// TIA Portal project "THELMA3_200224" (V15.1) (continued)
               #SDataDummy := CONCAT(IN1 := #SDataDummy, IN2 := 'BBD');
               #SDataDummy := CONCAT(IN1 := #SDataDummy, IN2 := #ExtDate);
               Strg_TO_Chars(Strg := #SDataDummy,
                             pChars := 1,
                             Cnt => #Dummy2,
                             Chars := #SData);
               #SData[15 + #LenDummy] := #End;
               #SLen := 15 + #LenDummy + 1;
               #RLen := 3;
               #Step := 0;
               #STrig := TRUE;
               #RdataTime := FALSE;
               #RdataAlarm := FALSE;
               #RdataBatch := FALSE;
               #RdataBBD := TRUE;
               #RdataLabel := FALSE;
               #Selected := FALSE;
           ELSIF #MarketRegCode <> '' AND #ExtDate <> '' THEN // print all on the second row
               #CommandHead := 'U'; //head for update user field
               #LenDummy := LEN(#MarketRegCode);
               #SDataDummy := CONCAT(IN1 := #CommandHead, IN2 := #SecondField);
               #SDataDummy := CONCAT(IN1 := #SDataDummy, IN2 := #NewLine);
               #SDataDummy := CONCAT(IN1 := #SDataDummy, IN2 := #MarketRegCode);
               #SDataDummy := CONCAT(IN1 := #SDataDummy, IN2 := 'BBD');
               #SDataDummy := CONCAT(IN1 := #SDataDummy, IN2 := #ExtDate);
               Strg_TO_Chars(Strg := #SDataDummy,
                             pChars := 1,
                             Cnt => #Dummy2,
                             Chars := #SData);
               #SData[21 + #LenDummy] := #End;
               #SLen := 21 + #LenDummy + 1;
               #RLen := 3;
               #Step := 0;
               #STrig := TRUE;
               #RdataTime := FALSE;
               #RdataAlarm := FALSE;
               #RdataBatch := FALSE;
               #RdataBBD := TRUE;
               #RdataLabel := FALSE;
               #Selected := FALSE;
           END_IF;
       ELSIF #Step =5 THEN
           //command for selecting the label
           #CommandHead := 'M'; //head for current status of the printer
           #SData[0] := #Start;
           IF #MDR_Flag = TRUE THEN //select the MDR layout 
               #SDataDummy := CONCAT(IN1 := #CommandHead, IN2 := #MDR_LabelName);
               Strg_TO_Chars(Strg := #SDataDummy,
                             pChars := 1,
                             Cnt => #Dummy2,
                             Chars := #SData);
               #SData[5] := #End;
               #RLen := 3;
               #SLen := 6;
           ELSE
               #LenLabel := LEN(#NMDR_LabelName);
               #SDataDummy := CONCAT(IN1 := #CommandHead, IN2 := #NMDR_LabelName);
               Strg_TO_Chars(Strg := #SDataDummy,
                             pChars := 1,
                             Cnt => #Dummy2,
                             Chars := #SData);
               #SData[2+#LenLabel] := #End;
               #RLen := 3;
               #SLen := 3+#LenLabel;
           END_IF;
           #STrig := TRUE;
           #Step := 0;
           #RdataAlarm := FALSE;
           #RdataTime := FALSE;
           #RdataBatch := FALSE;
           #RdataBBD := FALSE;
           #RdataLabel := TRUE;
       ELSE
           #STrig := FALSE;
       END_IF;
   END_REGION

   REGION Feedback
       // Statement section REGION
       //Expect to receive "ACT"
       IF #DataReceived = TRUE THEN
           #StartTNR := FALSE;
           IF #RdataTime = TRUE THEN //check for the feedback for the time command
               FOR #i := 0 TO 56 DO
                   #TimeReceivedData[#i] := #RData[#i];
               END_FOR;
               IF #TimeReceivedData[0] = 16#24 THEN
                   #TimeOK := TRUE;
                   #TimeReceivedData[0] := 16#30;//clear the buffer
               ELSE
                   #TimeOK := FALSE;
               END_IF;
               #RdataTime := FALSE;
           ELSIF #RdataAlarm = TRUE THEN//check for the feedback for the alarm command
               FOR #i := 0 TO 56 DO
                   #AlarmReceivedData[#i] := #RData[#i];
               END_FOR;
               IF #AlarmReceivedData[7] = 16#30  THEN
                   #AlarmCheck := TRUE;

                   FOR #i := 0 TO 8 DO
                       #PrinterAlarmStatus[#i] := #AlarmReceivedData[#i];//save the status data for processing
                   END_FOR;
                   #AlarmReceivedData[7] := 16#31;//clear the buffer
               ELSE
                   #AlarmCheck := FALSE;
               END_IF;
               #RdataAlarm := FALSE;
           ELSIF #RdataBatch = TRUE THEN//check for the feedback for the buffer command
               FOR #i := 0 TO 56 DO
                   #BatchReceivedData[#i] := #RData[#i];
               END_FOR;
               IF #BatchReceivedData[0] = 16#24 THEN
                   #BatchOK := TRUE;
                   #BatchReceivedData[0] := 16#30;//clear the buffer
               ELSE
                   #BatchOK := FALSE;
               END_IF;
               #RdataBatch := FALSE;
           ELSIF #RdataBBD = TRUE THEN//check for the feedback for the buffer command
               FOR #i := 0 TO 56 DO
                   #BBD_ReceivedData[#i] := #RData[#i];
               END_FOR;
               IF #BBD_ReceivedData[0] = 16#24 THEN
                   #BBD_OK := TRUE;
                   #BBD_ReceivedData[0] := 16#30;//clear the buffer
               ELSE
                   #BBD_OK := FALSE;
               END_IF;
               #RdataBBD := FALSE;
           ELSIF #RdataLabel = TRUE THEN//check for the feedback for the buffer command
               FOR #i := 0 TO 56 DO
                   #LabelReceivedData[#i] := #RData[#i];
               END_FOR;
               IF #LabelReceivedData[0] = 16#24 THEN
                   #LabelOK := TRUE;
                   #LabelReceivedData[0] := 16#30;//clear the buffer
               ELSE
                   #LabelOK := FALSE;
               END_IF;
               #RdataLabel := FALSE;
           END_IF;
       ELSIF #DataSent = TRUE THEN // command send noting received
           #StartTNR := TRUE;
           IF #RdataTime = TRUE THEN
               #TimeOK := FALSE;
           END_IF;
           IF #RdataAlarm = TRUE THEN
               #AlarmCheck := FALSE;
           END_IF;
           IF #RdataBatch = TRUE THEN
               #BatchOK := FALSE;
           END_IF;
           IF #RdataBBD = TRUE THEN
               #BBD_OK := FALSE;
           END_IF;
           IF #RdataLabel = TRUE THEN
               #LabelOK := FALSE;
           END_IF;
       END_IF;
   END_REGION

   REGION Sending
       // Send the batch number when it is changed or for reconnection
       #SelectingR(CLK:=#LabelSelecting);
       #ReconnectR(CLK := #ConnectionStatus);
       #MDR_R(CLK := #MDR_Flag);
       #MDR_F(CLK := #MDR_Flag);
       #BlockedR(CLK := #BlockedProduct);
       #BlockedF(CLK := #BlockedProduct);
       //select the label
       IF #MDR_F.Q = TRUE OR #MDR_R.Q = TRUE OR #SelectingR.Q = TRUE OR #ReconnectR.Q = TRUE OR #NLabelChanged = TRUE THEN
           #Step := 5; //selecting the label
           IF #MDR_Flag = TRUE THEN
               #Selected := TRUE; //send the first row
               #First := TRUE;////send the second row
           END_IF;
       END_IF;
       // set the step to 3 after label is selected (small delay to make sure that the label is loaded)
       #BatchAfterLabelT(IN := #Selected,
                         PT := T#2S);
       IF #BatchAfterLabelT.Q = TRUE THEN
           #Step := 3;
       END_IF;
       //send the update information
       // Send the updateble data when it is changed and step 4 is done
       IF (#PlainDataChanged = TRUE OR #BlockedR.Q = TRUE OR #BlockedF.Q = TRUE) AND #SelectingR.Q = FALSE THEN
           #Step := 3; //send plain data
           #Selected := FALSE;
           #First := TRUE;
       END_IF;
       //set the step to 4 after the first row is send
       #SecondAfterFirstT(IN:=#First,
                          PT:=T#4S);
       IF #SecondAfterFirstT.Q = TRUE THEN
           #Step := 4;
       END_IF;
       // Send time and alarm commands
       //every 10 minute synchronise time
       #TimeSynchT(IN := #TimeSynchEnable,
                  PT := #TimeSynchPeriod);
       IF #TimeSynchT.Q = TRUE THEN
           #Step := 1;
           #TimeSynchEnable := FALSE;
       ELSIF #ConnectionStatus = TRUE AND NOT (#MDR_F.Q= TRUE OR #MDR_R.Q =TRUE OR #SelectingR.Q = TRUE OR #ReconnectR.Q = TRUE OR #NLabelChanged = TRUE) AND NOT (#PlainDataChanged = TRUE OR #BlockedR.Q = TRUE OR #BlockedF.Q = TRUE) THEN
           #TimeSynchEnable := TRUE;
       ELSE
           #TimeSynchEnable := FALSE;
       END_IF;
       //every 5 minute check for alarm
       #AlarmCheckT(IN := #AlarmCheckEnable,
                   PT := #AlarmCheckPeriod + T#20MS);//+20ms to avoid conflict
       IF #AlarmCheckT.Q = TRUE THEN
           #Step := 2;
           #AlarmCheckEnable := FALSE;
       ELSIF #ConnectionStatus = TRUE AND NOT (#MDR_F.Q = TRUE OR #MDR_R.Q = TRUE OR #SelectingR.Q = TRUE OR #ReconnectR.Q = TRUE OR #NLabelChanged = TRUE) AND NOT(#PlainDataChanged = TRUE OR #BlockedR.Q = TRUE OR #BlockedF.Q = TRUE) THEN
           #AlarmCheckEnable := TRUE;
       ELSE
           #AlarmCheckEnable := FALSE;
       END_IF;
   END_REGION

   REGION send try
       //if not receiving feedback after 10ms send a commad again
       #NotReceiveT(IN := #StartTNR,
                   PT := #TimeNR,
                   Q => #SendAgainTrigger);
       IF #SendAgainTrigger = TRUE THEN
           #StartTNR := FALSE;
       END_IF;
   END_REGION
   (*
   REGION ConnReestablised
       // connection Re-Established Rotinue. It try 5 times to connect to the printer, if not succsess enable time out error
       #ConnAgainT(IN := #ReTry,
                  PT := T#5S);// time out for reconnection
       //try five times to connect
       #ConnTryCountC(CU := #ReTry,
                     R := #ConnectionStatus,
                     PV := 5,
                     Q => #TimeOutError);
   END_REGION
   *)
END_REGION
END_FUNCTION_BLOCK

FUNCTION_BLOCK "CON_PlainHandle"   // FB2, FBD
{ S7_Optimized_Access := 'TRUE' }
VERSION : 0.1
   VAR_INPUT
      Heartbeat : Bool;
      NewArtBaseFlag : String;
      NewMDR_Flag : String;
      NewBatchNum : String;
      NewArtBaseNum : UDInt;
      NewMarketRegCode : String;
      NewBBD : String;
   END_VAR
   VAR_OUTPUT
      Error : Bool;
      ActualBatchNumSTR : String;
      ActualArtBaseNumSTR : String;
      ActualMarketRegCodeSTR : String;
      ActualBBD_STR : String;
      HeartbeatToPlain : Bool;
   END_VAR
   VAR
      NewDataPlain : Bool;
      ActualMDR_FlagSTR : String;
      ActualArtBaseFlagSTR : String;
      ActualBatchNum : String;
      ActualArtBaseNum : UDInt;
      ActualMDR_Flag : Bool;
      ActualArtFlag : Bool;
      HeartbeatT : TON_TIME;
      PrintSecondRow : Bool;
      HeartbeatT_2 : TON_TIME;
      CountC : CTU_INT;
   END_VAR
   VAR_TEMP
      i : Int;
      NewBatchLen : UInt;
      Correction : Array[0..13] of Char;
      CorrectionSTR : String;
      TmpB1 : Bool;
      TmpB2 : Bool;
   END_VAR
   VAR CONSTANT
      BatchSize : UInt := 10;
   END_VAR
BEGIN

REGION Network 1 (SCL)
   REGION connection
       // check the heartbeat from MES-OPC
     #HeartbeatT(IN:=NOT(#Heartbeat),
                 PT:=T#30S);
     IF #HeartbeatT.Q = TRUE THEN
         #TmpB1 := TRUE;
       ELSE
           #TmpB1 := FALSE;
       END_IF;
       #HeartbeatT_2(IN:=#Heartbeat,
                     PT:=T#30S);
       IF #HeartbeatT_2.Q = TRUE THEN
           #TmpB2 := TRUE;
       ELSE
           #TmpB2 := FALSE;
       END_IF;
       IF #TmpB1 OR #TmpB2 THEN
           #Error := 1;
       ELSE
           #Error := 0;
       END_IF;

       //Send the Heartbeat to MES-OPC
       #CountC(CU:="Clock_1Hz",
               PV:=15,
               Q=>#HeartbeatToPlain);
       IF #CountC.CV > 29 THEN
           #CountC.CV := 0;
       END_IF;
   END_REGION
   REGION Flags
       // check for flags 
       IF #NewArtBaseFlag = 'Y' THEN
           #ActualArtFlag := TRUE;
       ELSE
           #ActualArtFlag := FALSE;
       END_IF;
       IF #NewMDR_Flag = 'Y' THEN
           #ActualMDR_Flag := TRUE;
       ELSE
           #ActualMDR_Flag := FALSE;
       END_IF;
   END_REGION

   REGION input changing
       // check for input number changing

       IF  #NewBatchNum <> #ActualBatchNum  OR  #NewArtBaseNum <> #ActualArtBaseNum OR #NewMarketRegCode <>#ActualMarketRegCodeSTR OR #NewBBD <> #ActualBBD_STR OR #NewArtBaseFlag <> #ActualArtBaseFlagSTR THEN
           #NewDataPlain := TRUE;
       ELSE
           #NewDataPlain := FALSE;
       END_IF;
       IF #NewBBD <> #ActualBBD_STR OR #NewMarketRegCode <> #ActualMarketRegCodeSTR THEN
           #PrintSecondRow := TRUE;
       ELSE
           #PrintSecondRow := FALSE;
       END_IF;
    //   IF #NewMDR_Flag <> #ActualMDR_FlagSTR THEN
    //       #MDR_FlagChange := TRUE;
   //    ELSE
   //        #MDR_FlagChange := FALSE;
   //    END_IF;
     //  IF #NewArtBaseFlag <> #ActualArtBaseFlagSTR THEN
     //      #ArtBaseFlagChange := TRUE;
     //  ELSE
    //       #ArtBaseFlagChange := FALSE;
    //   END_IF;
   END_REGION
   REGION assign plain data
       FOR #i := 0 TO 13 DO
           #Correction[#i] := '0';
       END_FOR;
       // Statement section REGION
       #ActualArtBaseNum := #NewArtBaseNum;
       #ActualMarketRegCodeSTR := #NewMarketRegCode;
       #ActualBatchNum := #NewBatchNum;
       #ActualBBD_STR := #NewBBD;
       #ActualMDR_FlagSTR := #NewMDR_Flag;
       #ActualArtBaseFlagSTR := #NewArtBaseFlag;
       //Actual Batch in 10 digits (3 factoryID+7 batch ID)
       #NewBatchLen := INT_TO_UINT(LEN(#NewBatchNum));
       IF #NewBatchLen < #BatchSize THEN
           Chars_TO_Strg(Chars := #Correction,
                         pChars := 0,
                         Cnt := (#BatchSize - #NewBatchLen),
                         Strg => #CorrectionSTR);
           #ActualBatchNumSTR := CONCAT(IN1 := #CorrectionSTR, IN2 := #NewBatchNum);
       ELSE
           #ActualBatchNumSTR := #NewBatchNum;
       END_IF;
     //Art base number
       VAL_STRG(IN := #NewArtBaseNum,
                SIZE := 0,
                PREC := 0,
                FORMAT := 0,
                P := 1,
                OUT => #ActualArtBaseNumSTR);
   END_REGION
END_REGION
END_FUNCTION_BLOCK

FUNCTION_BLOCK "ProgramReader"   // FB3, FBD
{ S7_Optimized_Access := 'TRUE' }
VERSION : 0.1
   VAR_INPUT
      Value : Array[0..9] of Char;
      MaterialNumber : UDInt;
      ReaderRead : Bool;
      ReaderNoRead : Bool;
      ExtTrigger : Bool;
      ResetFaults : Bool;
      ResetCounters : Bool;
   END_VAR
   VAR_OUTPUT
      Reading : UDInt;
      Msg_NoRead : Bool;
      Fault_MisMatch : Bool;
      Fault_NoRead : Bool;
      Fault_Trigger : Bool;
   END_VAR
   VAR_IN_OUT
      NumGross : UDInt;
      NumRead : UDInt;
      NumNoRead : UDInt;
      NumMatch : UDInt;
      NumNoMatch : UDInt;
   END_VAR
   VAR
      ReadingDInt : UDInt;
      ReadingSTR : String;
      MaterialNumberSTR : String;
      CompDINOut1 : Bool;
      HF_PosEdge1 : Bool;
      HF_PosEdge2 : Bool;
      HF_PosEdge3 : Bool;
      HF_PosEdge4 : Bool;
      HF_PosEdge5 : Bool;
      HF_PosEdge6 : Bool;
      HF_PosEdge7 : Bool;
      HF_PosEdge8 : Bool;
      HF_PosEdge9 : Bool;
      HF_NegEdge1 : Bool;
      HF_NegEdge2 : Bool;
      HF_MisMatch : Bool;
      HF_NoRead : Bool;
      HF_FltTrigger : Bool;
      HF_MisTrigger : Bool;
      HF_FltNoRead : Bool;
      T_FltNoRead : IEC_TIMER;
      Time_FltNoRead : Time := T#500MS;
      T_FltTriggerWatchdog : IEC_TIMER;
      Time_FltTriggerWatchdog : Time := T#5s;
   END_VAR
   VAR RETAIN
      C_FltNoRead : IEC_COUNTER;
      C_FltNoRead100 : IEC_COUNTER;
   END_VAR
   VAR
      TriggerCTR : "Counter_32Bit";
      ReadCTR : "Counter_32Bit";
      NoReadCTR : "Counter_32Bit";
      MatchCTR : "Counter_32Bit";
      NoMatchCTR : "Counter_32Bit";
      IEC_Timer_0_Instance : TP_TIME;
      MisTriggerCTR : "Counter_32Bit";
      NumMisTrigger : UDInt;
      NumNoReadGross : UDInt;
      EmptyBuffer : Bool;
      ReadData : Bool;
      DataValid : Bool;
      IEC_Timer_0_Instance_1 : TON_TIME;
   END_VAR
   VAR RETAIN
      Mis_3_row : CTU_INT;
   END_VAR
   VAR_TEMP   // added for the SCL form of the ladder/FBD networks
      _w1 : Bool;
   END_VAR
BEGIN

REGION Network 1
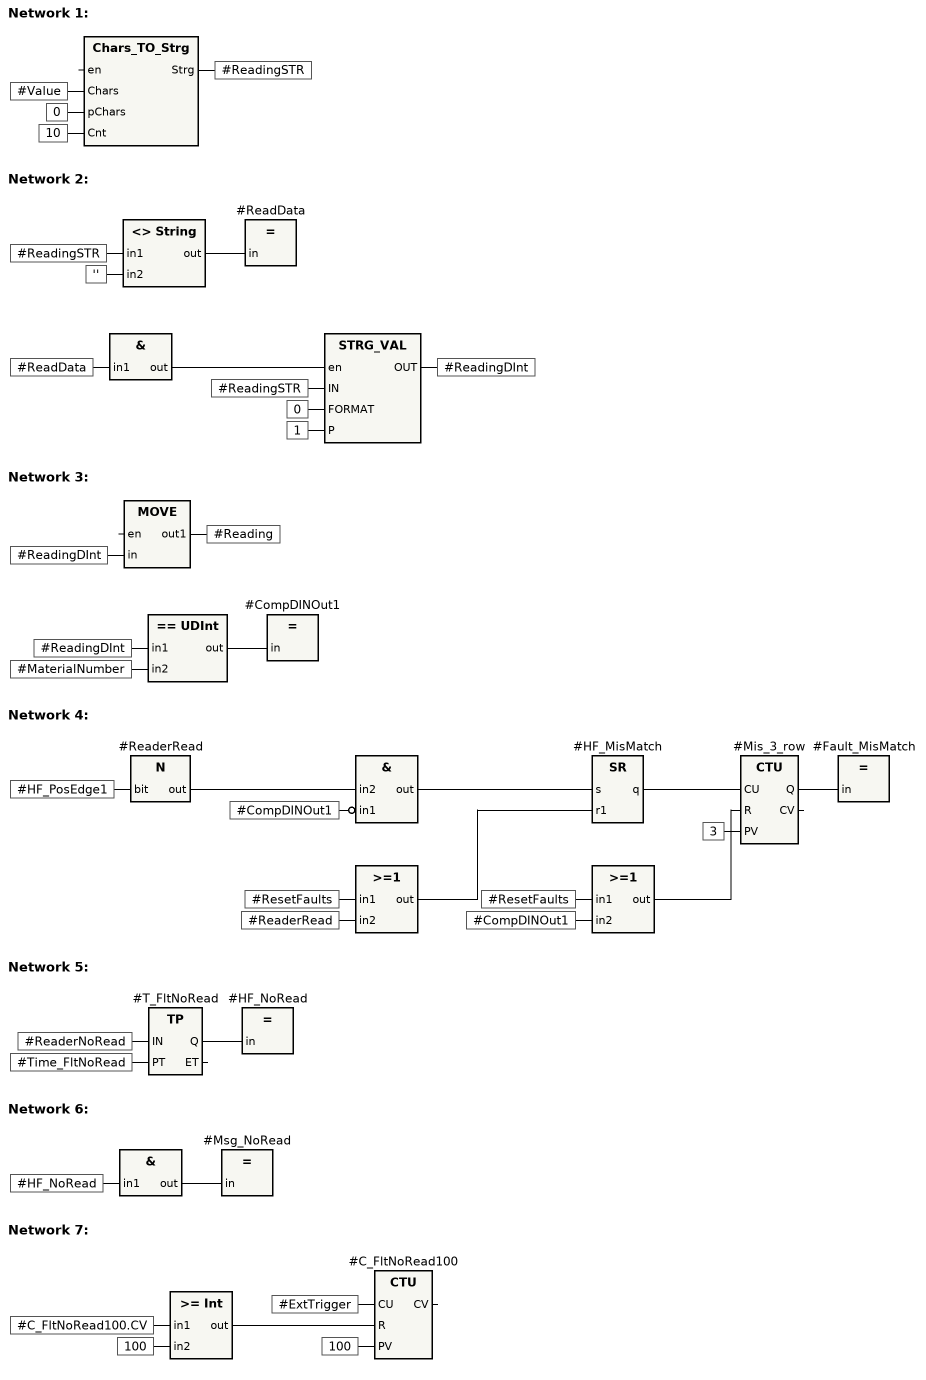
   // no SCL statement known for Chars_TO_Strg: written as a call
   Chars_TO_Strg(Chars := #Value, pChars := 0, Cnt := 10, Strg => #ReadingSTR);
END_REGION

REGION Network 2
   #ReadData := #ReadingSTR <> '';
   IF #ReadData THEN STRG_VAL(IN := #ReadingSTR, FORMAT := 0, P := 1, OUT => #ReadingDInt); END_IF;
END_REGION

REGION Network 3
   #Reading := #ReadingDInt;
   #CompDINOut1 := #ReadingDInt = #MaterialNumber;
END_REGION

REGION Network 4
   #_w1 := NOT #ReaderRead AND #HF_PosEdge1;   // falling edge of #ReaderRead
   #HF_PosEdge1 := #ReaderRead;
   IF #_w1 AND NOT #CompDINOut1 THEN
       #HF_MisMatch := TRUE;   // SR flip-flop
   END_IF;
   IF #ResetFaults OR #ReaderRead THEN #HF_MisMatch := FALSE; END_IF;
   #Mis_3_row(CU := #HF_MisMatch, R := #ResetFaults OR #CompDINOut1, PV := 3);   // CTU
   #Fault_MisMatch := #Mis_3_row.Q;
END_REGION

REGION Network 5
   #T_FltNoRead.TP(IN := #ReaderNoRead, PT := #Time_FltNoRead);
   #HF_NoRead := #T_FltNoRead.Q;
END_REGION

REGION Network 6
   #Msg_NoRead := #HF_NoRead;
END_REGION

REGION Network 7
   #C_FltNoRead100.CTU(CU := #ExtTrigger, R := #C_FltNoRead100.CV >= 100, PV := 100);
END_REGION

REGION Network 8
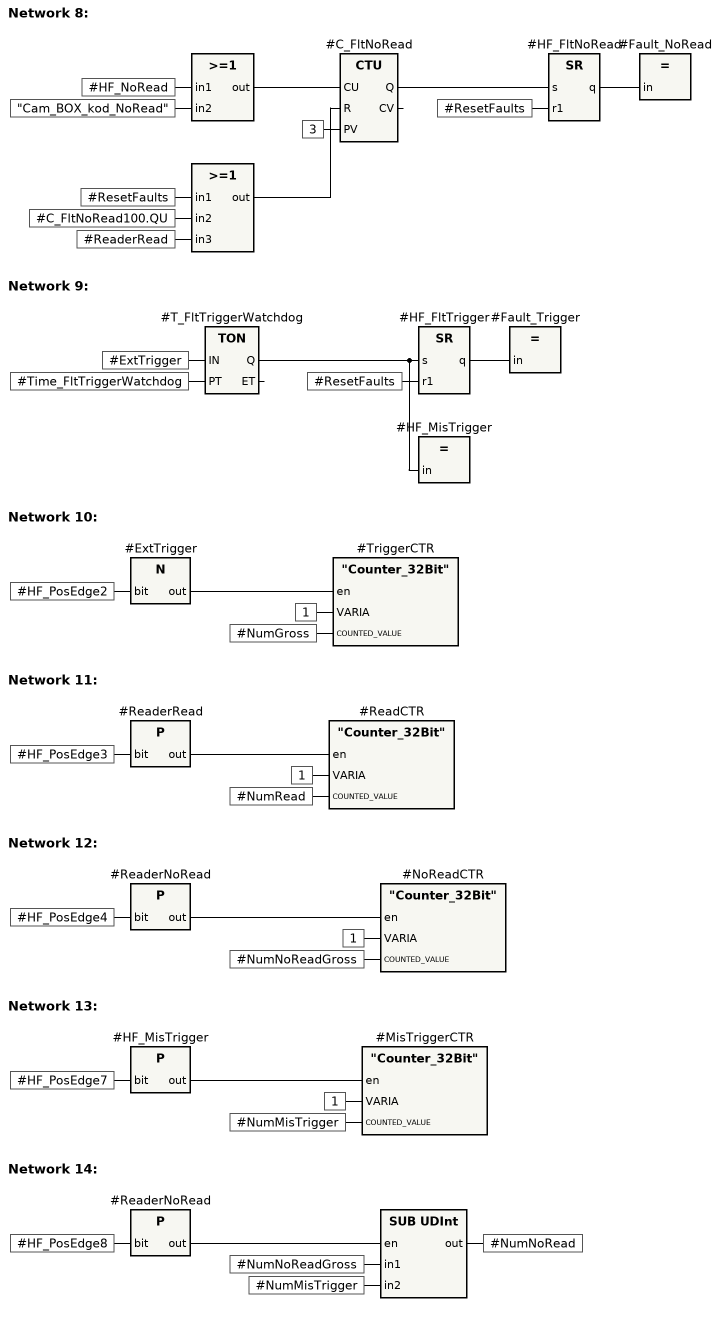
   #C_FltNoRead.CTU(CU := #HF_NoRead OR "Cam_BOX_kod_NoRead",
                    R := #ResetFaults OR #C_FltNoRead100.QU OR #ReaderRead,
                    PV := 3);
   IF #C_FltNoRead.Q THEN
       #HF_FltNoRead := TRUE;   // SR flip-flop
   END_IF;
   IF #ResetFaults THEN #HF_FltNoRead := FALSE; END_IF;
   #Fault_NoRead := #HF_FltNoRead;
END_REGION

REGION Network 9
   #T_FltTriggerWatchdog.TON(IN := #ExtTrigger, PT := #Time_FltTriggerWatchdog);
   IF #T_FltTriggerWatchdog.Q THEN
       #HF_FltTrigger := TRUE;   // SR flip-flop
   END_IF;
   IF #ResetFaults THEN #HF_FltTrigger := FALSE; END_IF;
   #Fault_Trigger := #HF_FltTrigger;
   #HF_MisTrigger := #T_FltTriggerWatchdog.Q;
END_REGION

REGION Network 10
   #_w1 := NOT #ExtTrigger AND #HF_PosEdge2;   // falling edge of #ExtTrigger
   #HF_PosEdge2 := #ExtTrigger;
   IF #_w1 THEN
       #TriggerCTR(VARIA := 1, COUNTED_VALUE := #NumGross);   // "Counter_32Bit"
   END_IF;
END_REGION

REGION Network 11
   #_w1 := #ReaderRead AND NOT #HF_PosEdge3;   // rising edge of #ReaderRead
   #HF_PosEdge3 := #ReaderRead;
   IF #_w1 THEN
       #ReadCTR(VARIA := 1, COUNTED_VALUE := #NumRead);   // "Counter_32Bit"
   END_IF;
END_REGION

REGION Network 12
   #_w1 := #ReaderNoRead AND NOT #HF_PosEdge4;   // rising edge of #ReaderNoRead
   #HF_PosEdge4 := #ReaderNoRead;
   IF #_w1 THEN
       #NoReadCTR(VARIA := 1, COUNTED_VALUE := #NumNoReadGross);   // "Counter_32Bit"
   END_IF;
END_REGION

REGION Network 13
   #_w1 := #HF_MisTrigger AND NOT #HF_PosEdge7;   // rising edge of #HF_MisTrigger
   #HF_PosEdge7 := #HF_MisTrigger;
   IF #_w1 THEN
       #MisTriggerCTR(VARIA := 1, COUNTED_VALUE := #NumMisTrigger);   // "Counter_32Bit"
   END_IF;
END_REGION

REGION Network 14
   #_w1 := #ReaderNoRead AND NOT #HF_PosEdge8;   // rising edge of #ReaderNoRead
   #HF_PosEdge8 := #ReaderNoRead;
   IF #_w1 THEN #NumNoRead := #NumNoReadGross - #NumMisTrigger; END_IF;
END_REGION

REGION Network 15
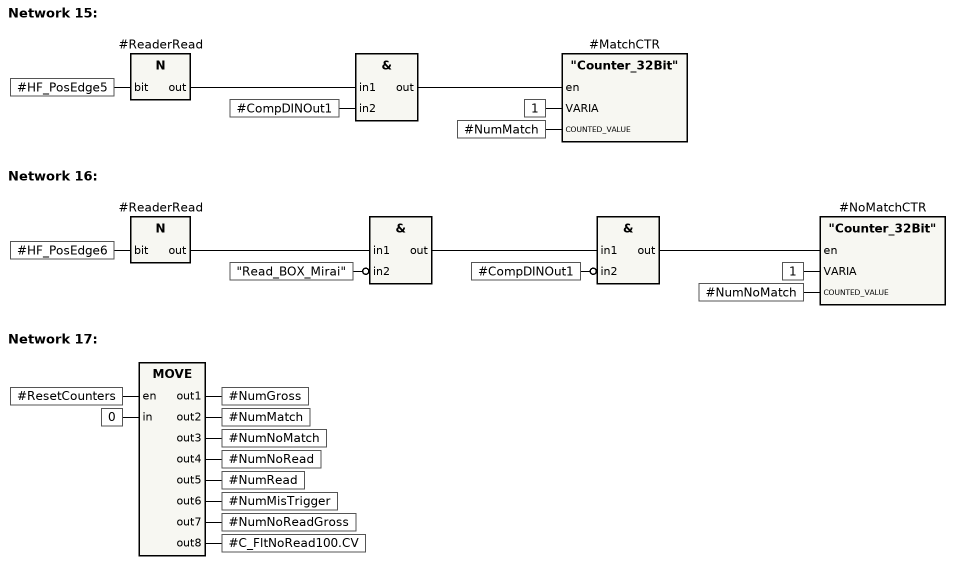
   #_w1 := NOT #ReaderRead AND #HF_PosEdge5;   // falling edge of #ReaderRead
   #HF_PosEdge5 := #ReaderRead;
   IF #_w1 AND #CompDINOut1 THEN
       #MatchCTR(VARIA := 1, COUNTED_VALUE := #NumMatch);   // "Counter_32Bit"
   END_IF;
END_REGION

REGION Network 16
   #_w1 := NOT #ReaderRead AND #HF_PosEdge6;   // falling edge of #ReaderRead
   #HF_PosEdge6 := #ReaderRead;
   IF #_w1 AND NOT "Read_BOX_Mirai" AND NOT #CompDINOut1 THEN
       #NoMatchCTR(VARIA := 1, COUNTED_VALUE := #NumNoMatch);   // "Counter_32Bit"
   END_IF;
END_REGION

REGION Network 17
   IF #ResetCounters THEN
       #NumGross := 0;
       #NumMatch := 0;
       #NumNoMatch := 0;
       #NumNoRead := 0;
       #NumRead := 0;
       #NumMisTrigger := 0;
       #NumNoReadGross := 0;
       #C_FltNoRead100.CV := 0;
   END_IF;
END_REGION
END_FUNCTION_BLOCK

FUNCTION_BLOCK "SimpleRead"   // FB4, FBD
{ S7_Optimized_Access := 'TRUE' }
VERSION : 0.1
   VAR_INPUT
      ExtTrigger : Bool := false;
      ResultAvailable : Bool;
      TriggerReady : Bool;
      TriggerAck : Bool;
      ResultID : Word;
      ResultCode : Word;
      ResultLength : Word;
      TriggerDelayTime : Time := T#10ms;
      SrcValue : ANY;
   END_VAR
   VAR_OUTPUT
      ID : Int;
      Flags : Int;
      Length : Int;
      TriggerEnable : Bool;
      TriggerReader : Bool;
      ResultsAck : Bool;
   END_VAR
   VAR_IN_OUT
      DstValue : ANY;
   END_VAR
   VAR
      ResultPending : Bool;
      Timer1 : IEC_TIMER;
      T_DelayTrigger : IEC_TIMER;
      HF_TriggerEnable : Bool;
      HF_TriggerReader : Bool;
      HF_ResultsAck : Bool;
      HF_DelayTrigger : Bool;
      IntTrigger : Bool;
   END_VAR
   VAR_TEMP
      BLKMOVRES : Int;
      Done : Bool;
   END_VAR
   VAR_TEMP   // added for the SCL form of the ladder/FBD networks
      _w1 : Bool;
   END_VAR
BEGIN

REGION Network 1
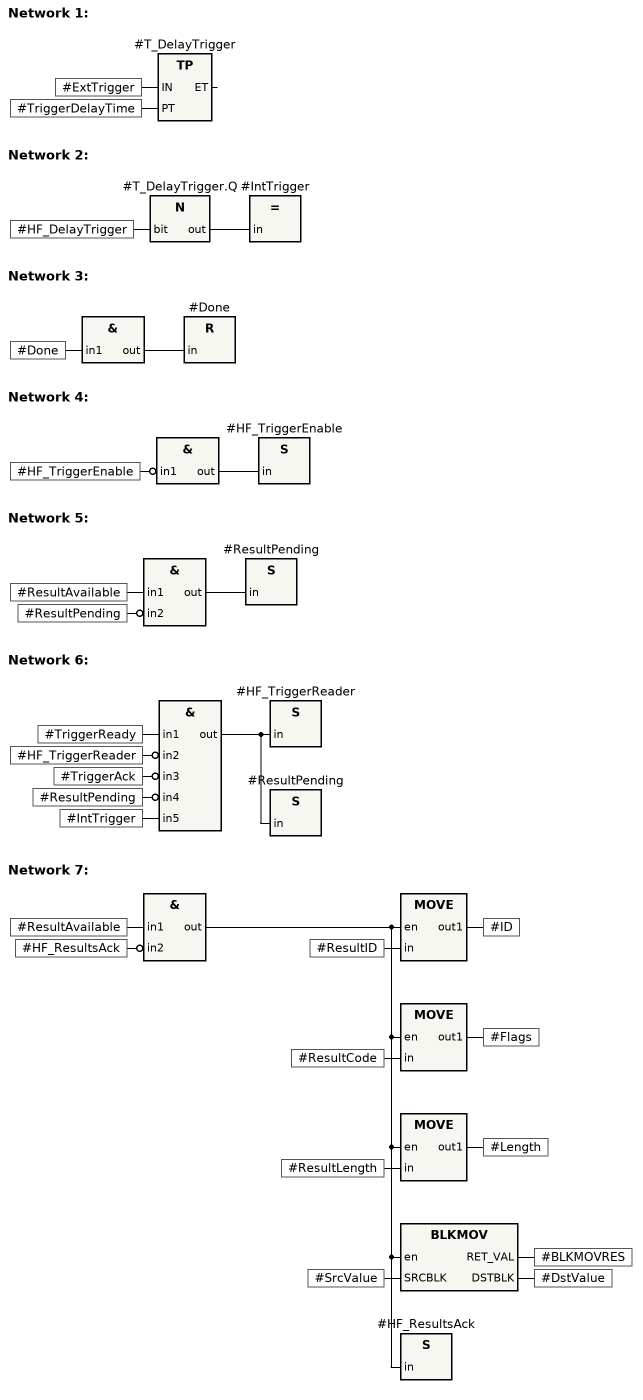
   #T_DelayTrigger.TP(IN := #ExtTrigger, PT := #TriggerDelayTime);
END_REGION

REGION Network 2
   #_w1 := NOT #T_DelayTrigger.Q AND #HF_DelayTrigger;   // falling edge of #T_DelayTrigger.Q
   #HF_DelayTrigger := #T_DelayTrigger.Q;
   #IntTrigger := #_w1;
END_REGION

REGION Network 3
   IF #Done THEN #Done := FALSE; END_IF;
END_REGION

REGION Network 4
   IF NOT #HF_TriggerEnable THEN #HF_TriggerEnable := TRUE; END_IF;
END_REGION

REGION Network 5
   IF #ResultAvailable AND NOT #ResultPending THEN #ResultPending := TRUE; END_IF;
END_REGION

REGION Network 6
   #_w1 := #TriggerReady AND NOT #HF_TriggerReader AND NOT #TriggerAck AND NOT #ResultPending AND #IntTrigger;
   IF #_w1 THEN
       #HF_TriggerReader := TRUE;
       #ResultPending := TRUE;
   END_IF;
END_REGION

REGION Network 7
   IF #ResultAvailable AND NOT #HF_ResultsAck THEN
       #ID := #ResultID;
       #Flags := #ResultCode;
       #Length := #ResultLength;
       #BLKMOVRES := BLKMOV(SRCBLK := #SrcValue, DSTBLK => #DstValue);
       #HF_ResultsAck := TRUE;
   END_IF;
END_REGION

REGION Network 8
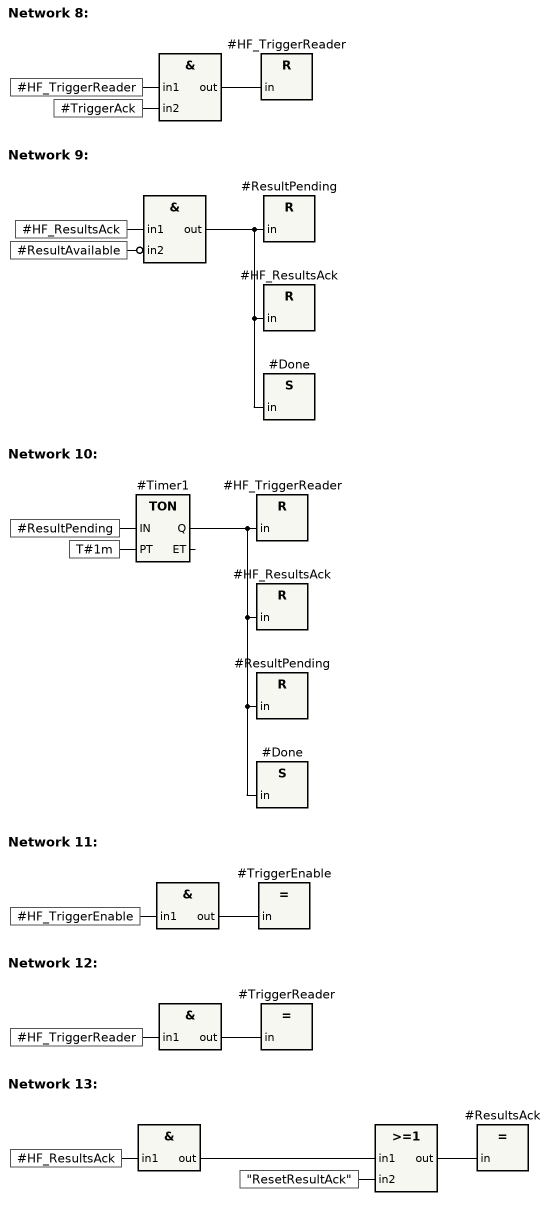
   IF #HF_TriggerReader AND #TriggerAck THEN #HF_TriggerReader := FALSE; END_IF;
END_REGION

REGION Network 9
   IF #HF_ResultsAck AND NOT #ResultAvailable THEN #ResultPending := FALSE; END_IF;
   #_w1 := #HF_ResultsAck AND NOT #ResultAvailable;
   IF #_w1 THEN
       #HF_ResultsAck := FALSE;
       #Done := TRUE;
   END_IF;
END_REGION

REGION Network 10
   #Timer1.TON(IN := #ResultPending, PT := T#1m);
   IF #Timer1.Q THEN
       #HF_TriggerReader := FALSE;
       #HF_ResultsAck := FALSE;
       #ResultPending := FALSE;
       #Done := TRUE;
   END_IF;
END_REGION

REGION Network 11
   #TriggerEnable := #HF_TriggerEnable;
END_REGION

REGION Network 12
   #TriggerReader := #HF_TriggerReader;
END_REGION

REGION Network 13
   #ResultsAck := #HF_ResultsAck OR "ResetResultAck";
END_REGION

REGION Network 14 (STL)
         A     #Done;
         SAVE;
END_REGION
END_FUNCTION_BLOCK

FUNCTION_BLOCK "MarkemImaje_2200"   // FB5, FBD
{ S7_Optimized_Access := 'TRUE' }
VERSION : 0.1
   VAR_INPUT
      RemoteAddress : String[20];
      ConnectionStatus : Bool;
      Inverse : Bool;
      LabelSelecting : Bool;
      ID : Conn_Ouc;
      ConType : Bool;
      BatchNumber : String;
      GTIN_Number : String;
      ArtNumber : String;
      MachineID : String;
      ExtDate : String;
      PlainDataChanged : Bool;
      "Date" : String;
      "Time" : String;
      DataReceived : Bool;
      DataSent : Bool;
      TimeSynchPeriod : Time := T#10M;
      AlarmCheckPeriod : Time := T#3M;
      RData : Array[0..56] of Byte;
      ExtTrigger : Bool;
      Stop : Bool;
   END_VAR
   VAR_OUTPUT
      Serial : UDInt;
      ErrorIP : Bool;
      BatchOK : Bool;
      AlarmCheck : Bool;
      TimeOK : Bool;
      LabelOK : Bool;
   END_VAR
   VAR
      Config : TADDR_Param;
      Configuration : "typeLCom_Config";
      RLen : UDInt;
      SLen : UDInt;
      SData : Array[0..95] of Byte;
      StartTNR : Bool;
      TimeNR : Time := T#1m;
      SendAgainTrigger : Bool;
      ExpFlag : Bool;
      NotReceiveT : TON_TIME;
      TimeSynchEnable : Bool := false;
      TimeSynchT : TON_TIME;
      AlarmCheckEnable : Bool := false;
      AlarmCheckT : TON_TIME;
      STrig : Bool;
      "Step" : UDInt;
      AlarmReceivedData : Array[0..56] of Byte;
      TimeReceivedData : Array[0..56] of Byte;
      BatchReceivedData : Array[0..56] of Byte;
      MacroReceivedData : Array[0..56] of Byte;
      RdataTime : Bool;
      RdataAlarm : Bool;
      RdataBatch : Bool;
      RdataMacro : Bool;
      DatePrinted : String;
      TimePrinted : String;
      DateChar : Array[0..7] of Char;
      TimeChar : Array[0..5] of Char;
      ReconnectR : R_TRIG;
      PrinterAlarmStatus : Array[0..31] of Bool;
      SelectingR : R_TRIG;
      Selected : Bool;
      InverseR : F_TRIG;
      InverseF : R_TRIG;
      ExtTriggerR : R_TRIG;
      SerialLen : Int;
      BatchAfterLabelT : TON_TIME;
      ChangeIP_T : TP_TIME;
      IP_Change : Bool;
      RemoteAddressOld : String;
   END_VAR
   VAR_TEMP
      StatusIP : Word;
      Dummy2 : UInt;
      i : Int;
      CommandHead : String;
      SerialSTR : String;
   END_VAR
   VAR CONSTANT
      Start : Char := '!';
      End : Char := '$R';
      NewLine : Char := '$L';
      LabelNameExp : String := 'EssityBBD___';
      LabelNameExpInv : String := 'EssityBBDInv';
      LabelName : String := 'Essity______';
      LabelNameInv : String := 'Essity___Inv';
   END_VAR
BEGIN

